// Mitsubishi GX Works2 project: Calculate   PLC: Q06UDEH

TYPE ConveyorIO : STRUCT
  xCWPresent : BOOL;  (* 正转检测有无传感器 *)
  xCCWPresent : BOOL;  (* 反转检测有无传感器 *)
  xLoad : BOOL;  (* 上料请求 *)
  xUnload : BOOL;  (* 下料请求 *)
  xMotorCW : BOOL;  (* 电机正转 *)
  xMotorCCW : BOOL;  (* 电机反转 *)
  xEmpty : BOOL;  (* 线体状态为空 *)
  xNextRun : BOOL;  (* 下段线体运行 *)
  xUnloadCCW : BOOL;  (* 下料为反转 *)
  xloadCCW : BOOL;  (* 上料为反转 *)
  xLeave : BOOL;  (* 已经离开 *)
  xForward : BOOL;  (* 正转手动 *)
  xBackward : BOOL;  (* 反转手动 *)
  xBusy : BOOL;  (* 工作中 *)
  xPutInto : BOOL;  (* 线体直接投入物料 *)
  xLoadAlarrm : BOOL;  (* 上料报警 *)
  xUnloadAlarm : BOOL;  (* 下料报警 *)
  iProductCategory : INT;  (* 产品种类 *)
  tLeaveDelay : TIME;  (* 离开延时设置 *)
  tLoadDelay : TIME;  (* 进入延时设置 *)
END_STRUCT END_TYPE

TYPE ShuttleCarIO : STRUCT
  xReady : BOOL;  (* 准备就绪 *)
  xForward : BOOL;  (* 正转 *)
  xBackward : BOOL;  (* 反转 *)
  iCurrentPos : INT;  (* 当前位置 *)
  iDestinationPos : INT;  (* 目标位置 *)
  xCW : BOOL;  (* 正转输出 *)
  xCCW : BOOL;  (* 反转输出 *)
  xBrake : BOOL;  (* 刹车 *)
  xHomeSwitch : BOOL;  (* 零位接近开关 *)
  xPosLimit : BOOL;  (* 正限位 *)
  xNegLimit : BOOL;  (* 负限位 *)
  xMDIExe : BOOL;  (* MDI开始 *)
  xMDIDone : BOOL;  (* MDI 完成 *)
  xPassLimit : BOOL;  (* 限位屏蔽 *)
  xPosLimitCatch : BOOL;  (* 正限位捕捉 *)
  xNegLimitCatch : BOOL;  (* 负限位捕捉 *)
  xHomeExe : BOOL;  (* 开始寻零 *)
  xHomeDone : BOOL;  (* 寻零完成 *)
  xHomeBusy : BOOL;  (* 寻零中 *)
  xHomeFailed : BOOL;  (* 寻零失败 *)
  xBusy : BOOL;  (* 工作中 *)
END_STRUCT END_TYPE

TYPE SwitchIO : STRUCT
  xLiftCylinderRetractDetect : BOOL;
  xLiftCylinderExtendDetect : BOOL;
  xLiftCylinderRetract : BOOL;
  xLiftCylinderExtend : BOOL;
  xEntryBarCylinderRetract : BOOL;
  xLiftCylinderExtendInit : BOOL;
  xEntryEnable : BOOL;
  xExitEnable : BOOL;
  xExitBarCylinderRetract : BOOL;
  xSwithEnable : BOOL;
  xLiftCylinderRetractButton : BOOL;
  xLiftCylinderExtendButton : BOOL;
  xEntryBarCylinderRetractButton : BOOL;
  xExitBarCylinderRetractButton : BOOL;
END_STRUCT END_TYPE

// global labels: Global1
VAR_GLOBAL
  g_xAuto : BOOL;
  g_xManual : BOOL;
  g_xEStop AT X23 : BOOL;
  g_xReset AT X20 : BOOL;
  g_xStackLampRed AT Y120 : BOOL;
  g_xStackLampAmber AT Y121 : BOOL;
  g_xStackLampGreen AT Y122 : BOOL;
  g_xBuzzer AT Y123 : BOOL;
  g_xStop AT M2 : BOOL;
  g_xLocalAutoStart AT M1 : BOOL;
  g_xRemoteAutoStart AT M0 : BOOL;
  g_xRemoteAuto AT M10 : BOOL;
  g_iState AT D40 : INT;
  g_iLocalAutoStep : INT;
END_VAR

// task Task_01 (event TRUE, interval 0, priority 31): POU, Start, UDP

PROGRAM POU
VAR
  H3000Conveyor1 : Conveyor;
  H3000Conveyor1IO : ConveyorIO;
  H3000Conveyor2 : Conveyor;
  H3000Conveyor2IO : ConveyorIO;
  H3000Conveyor3 : Conveyor;
  H3000Conveyor3IO : ConveyorIO;
  H3000Conveyor4 : Conveyor;
  H3000Conveyor4IO : ConveyorIO;
  H3000Conveyor5 : Conveyor;
  H3000Conveyor5IO : ConveyorIO;
  H3000Conveyor6 : Conveyor;
  H3000Conveyor6IO : ConveyorIO;
  H3000Conveyor7 : Conveyor;
  H3000Conveyor7IO : ConveyorIO;
  H3000Conveyor8 : Conveyor;
  H3000Conveyor8IO : ConveyorIO;
  H3000Conveyor9 : Conveyor;
  H3000Conveyor9IO : ConveyorIO;
  H3000Conveyor10 : Conveyor;
  H3000Conveyor10IO : ConveyorIO;
  H3000ChemConveyor1 : Conveyor;
  H3000ChemConveyor1IO : ConveyorIO;
  H3000ChemConveyor2 : Conveyor;
  H3000ChemConveyor2IO : ConveyorIO;
  H3000ChemConveyor3 : Conveyor;
  H3000ChemConveyor3IO : ConveyorIO;
  Lifter1 : ShuttleCar;
  Lifter1IO : ShuttleCarIO;
  Conveyor1 : Conveyor;
  Conveyor1IO : ConveyorIO;
  Lifter2 : ShuttleCar;
  Lifter2IO : ShuttleCarIO;
  Conveyor2 : Conveyor;
  Conveyor2IO : ConveyorIO;
  H2200Conveyor1 : Conveyor;
  H2200Conveyor1IO : ConveyorIO;
  H2200Conveyor2 : Conveyor;
  H2200Conveyor2IO : ConveyorIO;
  H2200Conveyor3 : Conveyor;
  H2200Conveyor3IO : ConveyorIO;
  H2200Conveyor4 : Conveyor;
  H2200Conveyor4IO : ConveyorIO;
  H2200Conveyor5 : Conveyor;
  H2200Conveyor5IO : ConveyorIO;
  H2200Conveyor6 : Conveyor;
  H2200Conveyor6IO : ConveyorIO;
  H2200Conveyor7 : Conveyor;
  H2200Conveyor7IO : ConveyorIO;
  H2200Conveyor8 : Conveyor;
  H2200Conveyor8IO : ConveyorIO;
  H2200Conveyor9 : Conveyor;
  H2200Conveyor9IO : ConveyorIO;
  H2200Conveyor10 : Conveyor;
  H2200Conveyor10IO : ConveyorIO;
  H1000Conveyor1 : Conveyor;
  H1000Conveyor1IO : ConveyorIO;
  H1000Conveyor2 : Conveyor;
  H1000Conveyor2IO : ConveyorIO;
  H1000Conveyor3 : Conveyor;
  H1000Conveyor3IO : ConveyorIO;
  H1000Conveyor4 : Conveyor;
  H1000Conveyor4IO : ConveyorIO;
  H1000Conveyor5 : Conveyor;
  H1000Conveyor5IO : ConveyorIO;
  H1000Conveyor6 : Conveyor;
  H1000Conveyor6IO : ConveyorIO;
  H1000Conveyor7 : Conveyor;
  H1000Conveyor7IO : ConveyorIO;
  H1000Conveyor8 : Conveyor;
  H1000Conveyor8IO : ConveyorIO;
  H1000Conveyor9 : Conveyor;
  H1000Conveyor9IO : ConveyorIO;
  H3000SwitchChem : Switch;
  H3000SwitchChemIO : SwitchIO;
  H850Switch : Switch;
  H850SwitchIO : SwitchIO;
  H850SwitchConveyorIn : ConveyorIO;
  H850SwitchConveyorOut : ConveyorIO;
  H850Conveyor8 : Conveyor;
  H850Conveyor8IO : ConveyorIO;
  H1000Conveyor10 : Conveyor;
  H1000Conveyor10IO : ConveyorIO;
  H3000SwitchChemConveyorIn : ConveyorIO;
  H3000SwitchChemConveyorOut : ConveyorIO;
  H3000SwitchQuadPackage : Switch;
  H3000SwitchQuadPackageIO : SwitchIO;
  H3000SwitchPackageConveyorIn : ConveyorIO;
  H3000SwitchPackageConveyorOut : ConveyorIO;
  H2200Switch1 : Switch;
  H2200Switch1IO : SwitchIO;
  H2200Switch1ConveyorIn : ConveyorIO;
  H2200Switch1ConveyorOut : ConveyorIO;
  H2200Switch2 : Switch;
  H2200Switch2IO : SwitchIO;
  H2200Switch2ConveyorIn : ConveyorIO;
  H2200Switch2ConveyorOut : ConveyorIO;
  iStep : INT;
  Import1Conveyor1 : Conveyor;
  Import1Conveyor1IO : ConveyorIO;
  Import1Conveyor2 : Conveyor;
  Import1Conveyor2IO : ConveyorIO;
  Import2Conveyor1 : Conveyor;
  Import2Conveyor1IO : ConveyorIO;
  Import2Conveyor2 : Conveyor;
  Import2Conveyor2IO : ConveyorIO;
  Export1Conveyor1 : Conveyor;
  Export1Conveyor1IO : ConveyorIO;
  Export1Conveyor2 : Conveyor;
  Export1Conveyor2IO : ConveyorIO;
  Export2Conveyor1 : Conveyor;
  Export2Conveyor1IO : ConveyorIO;
  Export2Conveyor2 : Conveyor;
  Export2Conveyor2IO : ConveyorIO;
  Export2Switch : Switch;
  Export2SwitchIO : SwitchIO;
  Export2SwitchConveyorIn : ConveyorIO;
  Export2SwitchConveyorOut : ConveyorIO;
  H850Rotor : ShuttleCar;
  H850RotorIO : ShuttleCarIO;
  H850RotorConveyor : Conveyor;
  H850RotorConveyorIO : ConveyorIO;
  H2200RotorIO : ShuttleCarIO;
  H2200RotorConveyor : Conveyor;
  H2200RotorConveyorIO : ConveyorIO;
  H2200Rotor : ShuttleCar;
  H850Conveyor1 : Conveyor;
  H850Conveyor1IO : ConveyorIO;
  H850Conveyor3 : Conveyor;
  H850Conveyor3IO : ConveyorIO;
  H850Conveyor4 : Conveyor;
  H850Conveyor4IO : ConveyorIO;
  H850Conveyor5 : Conveyor;
  H850Conveyor5IO : ConveyorIO;
  H850Conveyor6 : Conveyor;
  H850Conveyor6IO : ConveyorIO;
  Lifter2Position : ARRAY [0..5] OF INT;
  ii : INT;
  H2200SwitchEmptyABack : Switch;
  H2200SwitchEmptyABackIO : SwitchIO;
  H2200SwitchEmptyABackConveyorIn : ConveyorIO;
  H2200SwitchEmptyABackConveyorOut : ConveyorIO;
  H2200SwitchEmptyBBack : Switch;
  H2200SwitchEmptyBBackIO : SwitchIO;
  H2200SwitchEmptyBBackConveyorIn : ConveyorIO;
  H2200SwitchEmptyBBackConveyorOut : ConveyorIO;
  H2200ImportConveyor1 : Conveyor;
  H2200ImportConveyor1IO : ConveyorIO;
  H2200ImportConveyor2 : Conveyor;
  H2200ImportConveyor2IO : ConveyorIO;
  Import1Switch : Switch;
  Import1SwitchIO : SwitchIO;
  Import1SwitchConveyorIn : ConveyorIO;
  Import1SwitchConveyorOut : ConveyorIO;
  Export1Switch : Switch;
  Export1SwitchIO : SwitchIO;
  Export1SwitchConveyorIn : ConveyorIO;
  Export1SwitchConveyorOut : ConveyorIO;
  Import2Switch : Switch;
  Import2SwitchIO : SwitchIO;
  Import2SwitchConveyorIn : ConveyorIO;
  Import2SwitchConveyorOut : ConveyorIO;
  Import1LoadCylinder : ShuttleCar;
  Import1LoadCylinderIO : ShuttleCarIO;
  Import2LoadCylinder : ShuttleCar;
  Import2LoadCylinderIO : ShuttleCarIO;
  Export1LoadCylinder : ShuttleCar;
  Export1LoadCylinderIO : ShuttleCarIO;
  Export2LoadCylinder : ShuttleCar;
  Export2LoadCylinderIO : ShuttleCarIO;
  Lifter2Occupy : BOOL;  (* 提升机2占用标志位 *)
  Lifter2ChemImport : BOOL;  (* 提升机2化成入库 *)
  Lifter2ExportChem : BOOL;  (* 提升机2出库到化成 *)
END_VAR
H3000SwitchQuadPackage(ConveyorEntryIO:=H3000SwitchPackageConveyorIn ,
                                                        ConveyorExitIO:=H3000SwitchPackageConveyorOut ,
                                                        SwitchIO:=H3000SwitchQuadPackageIO );
H3000SwitchQuadPackageIO.xLiftCylinderExtendButton:=M75;
H3000SwitchQuadPackageIO.xLiftCylinderRetractButton:=M76;
H3000SwitchQuadPackageIO.xExitBarCylinderRetractButton:=M83;
Y128:=H3000SwitchQuadPackageIO.xEXITBarCylinderRetract;
Y12C:=H3000SwitchQuadPackageIO.xLiftCylinderExtend;
Y12A:=H3000SwitchQuadPackageIO.xLiftCylinderRetract;
H3000SwitchQuadPackageIO.xLiftCylinderExtendDetect:=X29;
H3000SwitchQuadPackageIO.xLiftCylinderRetractDetect:=X2A;
H3000SwitchPackageConveyorIn.xForward:=M77;
H3000SwitchPackageConveyorIn.xCWPresent:=X28;
(*Y187:=H3000SwitchPackageConveyorIn.xMotorCW;*)
H3000SwitchPackageConveyorOut.xForward:=M78;
H3000SwitchPackageConveyorOut.xCWPresent:=X2B;
Y12B:=H3000SwitchPackageConveyorOut.xMotorCW;

H3000SwitchChem(ConveyorEntryIO:=H3000SwitchChemConveyorIn ,
                                                        ConveyorExitIO:=H3000SwitchChemConveyorOut ,
                                                        SwitchIO:=H3000SwitchChemIO );
H3000SwitchChemIO.xLiftCylinderExtendButton:=M79;
H3000SwitchChemIO.xLiftCylinderRetractButton:=M80;
Y129:=H3000SwitchChemIO.xLiftCylinderExtend;
Y12D:=H3000SwitchChemIO.xLiftCylinderRetract;
H3000SwitchChemIO.xLiftCylinderExtendDetect:=X2C;
H3000SwitchChemIO.xLiftCylinderRetractDetect:=X2D;
H3000SwitchChemConveyorIn.xForward:=M81;
H3000SwitchChemConveyorIn.xCWPresent:=X2E;
Y19B:=H3000SwitchPackageConveyorIn.xMotorCW;
H3000SwitchChemConveyorOut.xForward:=M82;
H3000SwitchChemConveyorOut.xCWPresent:=X2E;
Y12E:=H3000SwitchChemConveyorOut.xMotorCW;
H3000SwitchChemIO.xSwithEnable:=1;

Lifter1(ShuttleCarInOut:=Lifter1IO);
ShuttleCarCurrentPosition( X8C OR X8D ,X8C ,X8D, FALSE, Lifter1IO.iCurrentPos );
Lifter1IO.xReady:=X24;
Lifter1Io.xForward:=M50 OR X91;
Lifter1IO.xBackward:=M51 OR X92;
Lifter1IO.xPosLimit:=X8E;
Lifter1IO.xNegLimit:=X8F;
Y18D:=Lifter1IO.xCW;
Y18E:=Lifter1IO.xCCW;
Y192:=Lifter1IO.xBrake;

Conveyor1(ConveyorMotor:=Conveyor1IO);
Conveyor1IO.xForward:=M52;
Conveyor1IO.xBackward:=M53;
Conveyor1IO.xCWPresent:=X93;
Conveyor1IO.xCCWPresent:=X94;
Y18B:=Conveyor1IO.xMotorCW;
Y18C:=Conveyor1IO.xMotorCCW;

Lifter2(ShuttleCarInOut:=Lifter2IO);
Lifter2Position[0]:=0;
Lifter2Position[1]:=57;
Lifter2Position[2]:=590;
Lifter2Position[3]:=5828;
Lifter2Position[4]:=6202;
Lifter2Position[5]:=9200;
FOR ii:=0 TO 5 BY 1 DO
	IF abs(D190-Lifter2Position[ii])<5 THEN
		Lifter2IO.iCurrentPos:=ii;
	END_IF;
END_FOR;
Lifter2IO.xReady:=X25;
(*提升机占用标志位控制*)
IF LIfter2IO.xBusy AND Conveyor2IO.xEmpty=0 AND g_xAuto THEN
	Lifter2Occupy:=1;
END_IF;
IF g_xManual OR g_xReset THEN
	Lifter2Occupy:=0;
END_IF;
IF ( Lifter2IO.iCurrentPos=1 AND NOT H850Conveyor8IO.xEmpty)   (*注液入库*)
	OR (Lifter2IO.iCurrentPos=2 AND NOT H1000Conveyor1IO.xEmpty)  (*化成入库*)
	OR (Lifter2IO.iCurrentPos=5  AND NOT H3000ChemConveyor3IO.xEmpty) THEN(*出库化成或空框去注液*)
	Lifter2Occupy:=1;
END_IF;
IF  (Lifter2IO.iCurrentPos=3 OR Lifter2IO.iCurrentPos=4) AND Conveyor2IO.xEmpty  THEN
	Lifter2Occupy:=0;
END_IF;

Lifter2Io.xForward:=M54 OR X9B;
Lifter2IO.xBackward:=M55 OR X9C;
Lifter2IO.xPosLimit:=X98;
Lifter2IO.xNegLimit:=X99;
Y193:=Lifter2IO.xCW;
Y194:=Lifter2IO.xCCW;
Y198:=Lifter2IO.xBrake;
(*提升机2编码器清零，到达负限位后清零*)
IF NOT Lifter2IO.xNegLimit THEN
	Y125:=1;
ELSE
	Y125:=0;
END_IF;

Conveyor2(ConveyorMotor:=Conveyor2IO);
Conveyor2IO.xForward:=M56;
Conveyor2IO.xBackward:=M57;
Conveyor2IO.xCWPresent:=X9D;
Conveyor2IO.xCCWPresent:=X9E;
Y19A:=Conveyor2IO.xMotorCW;
Y199:=Conveyor2IO.xMotorCCW;


H3000Conveyor1(ConveyorMotor:=H3000Conveyor1IO);
H3000Conveyor1IO.xForward:=M30;
H3000Conveyor1IO.xCWPresent:=X2F;
Y12F:=H3000Conveyor1IO.xMotorCW;

H3000Conveyor2(ConveyorMotor:=H3000Conveyor2IO);
H3000Conveyor2IO.xForward:=M31;
H3000Conveyor2IO.xCWPresent:=X30;
Y130:=H3000Conveyor2IO.xMotorCW;

H3000Conveyor3(ConveyorMotor:=H3000Conveyor3IO);
H3000Conveyor3IO.xForward:=M32;
H3000Conveyor3IO.xCWPresent:=X31;
Y131:=H3000Conveyor3IO.xMotorCW;

H3000Conveyor4(ConveyorMotor:=H3000Conveyor4IO);
H3000Conveyor4IO.xForward:=M33;
H3000Conveyor4IO.xCWPresent:=X32;
Y132:=H3000Conveyor4IO.xMotorCW;

H3000Conveyor5(ConveyorMotor:=H3000Conveyor5IO);
H3000Conveyor5IO.xForward:=M34;
H3000Conveyor5IO.xCWPresent:=X33;
Y133:=H3000Conveyor5IO.xMotorCW;

H3000Conveyor6(ConveyorMotor:=H3000Conveyor6IO);
H3000Conveyor6IO.xForward:=M34;
H3000Conveyor6IO.xCWPresent:=X34;
Y134:=H3000Conveyor6IO.xMotorCW;

H3000Conveyor7(ConveyorMotor:=H3000Conveyor7IO);
H3000Conveyor7IO.xForward:=M35;
H3000Conveyor7IO.xCWPresent:=X35;
Y135:=H3000Conveyor7IO.xMotorCW;
H3000Conveyor8(ConveyorMotor:=H3000Conveyor8IO);
H3000Conveyor8IO.xForward:=M36;
H3000Conveyor8IO.xCWPresent:=X36;
Y136:=H3000Conveyor8IO.xMotorCW;

H3000Conveyor9(ConveyorMotor:=H3000Conveyor9IO);
H3000Conveyor9IO.xForward:=M37;
H3000Conveyor9IO.xCWPresent:=X37;
Y137:=H3000Conveyor9IO.xMotorCW;

H3000Conveyor10(ConveyorMotor:=H3000Conveyor10IO);
H3000Conveyor10IO.xForward:=M38;
H3000Conveyor10IO.xCWPresent:=X38;
Y138:=H3000Conveyor10IO.xMotorCW;

H3000ChemConveyor1(ConveyorMotor:=H3000ChemConveyor1IO);
H3000ChemConveyor1IO.xForward:=M39;
H3000ChemConveyor1IO.xCWPresent:=X39;
Y139:=H3000ChemConveyor1IO.xMotorCW;

H3000ChemConveyor2(ConveyorMotor:=H3000ChemConveyor2IO);
H3000ChemConveyor2IO.xForward:=M40;
H3000ChemConveyor2IO.xCWPresent:=X3A;
Y13A:=H3000ChemConveyor2IO.xMotorCW;

H3000ChemConveyor3(ConveyorMotor:=H3000ChemConveyor3IO);
H3000ChemConveyor3IO.xForward:=M41;
H3000ChemConveyor3IO.xCWPresent:=X3B;
Y13B:=H3000ChemConveyor3IO.xMotorCW;

H2200Switch1(ConveyorEntryIO:=H2200Switch1ConveyorIn ,
                                                        ConveyorExitIO:=H2200Switch1ConveyorOut ,
                                                        SwitchIO:=H2200Switch1IO );
H2200Switch1IO.xLiftCylinderExtendButton:=M84;
H2200Switch1IO.xLiftCylinderRetractButton:=M85;
H2200Switch1IO.xExitBarCylinderRetractButton:=M86;
Y158:=H2200Switch1IO.xEXITBarCylinderRetract;
Y155:=H2200Switch1IO.xLiftCylinderExtend;
Y156:=H2200Switch1IO.xLiftCylinderRetract;
H2200Switch1IO.xLiftCylinderExtendDetect:=X55;
H2200Switch1IO.xLiftCylinderRetractDetect:=X56;
H2200Switch1ConveyorIn.xForward:=M87;
H2200Switch1ConveyorIn.xCWPresent:=X57;
Y177:=H2200Switch1ConveyorIn.xMotorCW;
H2200Switch1ConveyorOut .xForward:=M88;
H2200Switch1ConveyorOut .xCWPresent:=X57;
H2200Switch1ConveyorOut.tLoadDelay:=T#1s;
Y157:=H2200Switch1ConveyorOut .xMotorCW;

H2200ImportConveyor1(ConveyorMotor:=H2200ImportConveyor1IO);
H2200ImportConveyor1IO.xForward:=M136;
H2200ImportConveyor1IO.xCWPresent:=X53;
Y153:=H2200ImportConveyor1IO.xMotorCW;
H2200ImportConveyor2IO.tLeaveDelay:=T#5s;

H2200ImportConveyor2(ConveyorMotor:=H2200ImportConveyor2IO);
H2200ImportConveyor2IO.xForward:=M122;
H2200ImportConveyor2IO.xCWPresent:=X58;
Y154:=H2200ImportConveyor2IO.xMotorCW;
H2200ImportConveyor2IO.tLeaveDelay:=T#5s;

H2200Switch2(ConveyorEntryIO:=H2200Switch2ConveyorIn ,
                                                        ConveyorExitIO:=H2200Switch2ConveyorOut ,
                                                        SwitchIO:=H2200Switch2IO );
H2200Switch2IO.xLiftCylinderExtendButton:=M89;
H2200Switch2IO.xLiftCylinderRetractButton:=M90;
H2200Switch2IO.xExitBarCylinderRetractButton:=M91;
Y15C:=H2200Switch2IO.xEXITBarCylinderRetract;
Y159:=H2200Switch2IO.xLiftCylinderExtend;
Y15A:=H2200Switch2IO.xLiftCylinderRetract;
H2200Switch2IO.xLiftCylinderExtendDetect:=X59;
H2200Switch2IO.xLiftCylinderRetractDetect:=X5A;
H2200Switch2ConveyorIn.xForward:=M92;
H2200Switch2ConveyorIn.xCWPresent:=X5B;
H2200Switch2ConveyorIn.tLoadDelay:=T#2s;
Y15B:=H2200Switch2ConveyorIn.xMotorCW;
H2200Switch2ConveyorOut .xForward:=M93;
H2200Switch2ConveyorOut .xCWPresent:=X5B;
H2200Switch2ConveyorOut.tLeaveDelay:=T#8S;
H2200Switch2IO.xLiftCylinderExtendInit:=1;

H2200SwitchEmptyABack(ConveyorEntryIO:=H2200SwitchEmptyABackConveyorIn ,
                                                        ConveyorExitIO:=H2200SwitchEmptyABackConveyorOut ,
                                                        SwitchIO:=H2200SwitchEmptyABackIO );
H2200SwitchEmptyABackIO.xLiftCylinderExtendButton:=M137;
H2200SwitchEmptyABackIO.xLiftCylinderRetractButton:=M138;
H2200SwitchEmptyABackIO.xExitBarCylinderRetractButton:=M139;
Y160:=H2200SwitchEmptyABackIO.xLiftCylinderExtend;
Y161:=H2200SwitchEmptyABackIO.xLiftCylinderRetract;
H2200SwitchEmptyABackIO.xLiftCylinderExtendDetect:=X60;
H2200SwitchEmptyABackIO.xLiftCylinderRetractDetect:=X61;
H2200SwitchEmptyABackConveyorIn.xForward:=M140;
H2200SwitchEmptyABackConveyorIn.xCWPresent:=X62;
H2200SwitchEmptyABackConveyorIn.tLoadDelay:=T#2s;
Y162:=H2200SwitchEmptyABackConveyorIn.xMotorCW;
H2200SwitchEmptyABackConveyorOut .xForward:=M146;
H2200SwitchEmptyABackConveyorOut.xCWPresent:=X62;
H2200SwitchEmptyABackConveyorOut.tLeaveDelay:=T#30S;
Y177:=H2200SwitchEmptyABackConveyorOut .xMotorCW OR H2200SwitchEmptyBBackConveyorOut .xMotorCW ;

H2200SwitchEmptyBBack(ConveyorEntryIO:=H2200SwitchEmptyBBackConveyorIn ,
                                                        ConveyorExitIO:=H2200SwitchEmptyBBackConveyorOut ,
                                                        SwitchIO:=H2200SwitchEmptyBBackIO );
H2200SwitchEmptyBBackIO.xLiftCylinderExtendButton:=M141;
H2200SwitchEmptyBBackIO.xLiftCylinderRetractButton:=M142;
H2200SwitchEmptyBBackIO.xExitBarCylinderRetractButton:=M143;
Y166:=H2200SwitchEmptyBBackIO.xLiftCylinderExtend;
Y167:=H2200SwitchEmptyBBackIO.xLiftCylinderRetract;
H2200SwitchEmptyBBackIO.xLiftCylinderExtendDetect:=X66;
H2200SwitchEmptyBBackIO.xLiftCylinderRetractDetect:=X67;
H2200SwitchEmptyBBackConveyorIn.xForward:=M144;
H2200SwitchEmptyBBackConveyorIn.xCWPresent:=X68;
H2200SwitchEmptyBBackConveyorIn.tLoadDelay:=T#2s;
Y168:=H2200SwitchEmptyBBackConveyorIn.xMotorCW;
H2200SwitchEmptyBBackConveyorOut .xForward:=M145;
H2200SwitchEmptyBBackConveyorOut.xCWPresent:=X68;
H2200SwitchEmptyBBackConveyorOut.tLeaveDelay:=T#30S;

H2200Rotor(ShuttleCarInOut:=H2200RotorIO);
ShuttleCarCurrentPosition( X6F OR X75 ,X6F ,X75, FALSE, H2200RotorIO.iCurrentPos );
H2200RotorIO.xReady:=TRUE;
H2200RotorIO.xForward:=M78;
H2200RotorIO.xBackward:=M79;
H2200RotorIO.xPosLimit:=X71;
H2200RotorIO.xNegLimit:=X72;
Y170:=H2200RotorIO.xCW;
Y16F:=H2200RotorIO.xCCW;
Y1B8:=H2200RotorIO.xBrake;

H2200RotorConveyor(ConveyorMotor:=H2200RotorConveyorIO);
H2200RotorConveyorIO.xForward:=M80;
H2200RotorConveyorIO.xBackward:=M81;
H2200RotorConveyorIO.xCWPresent:=X74;
H2200RotorConveyorIO.xCcWPresent:=X73;
Y172:=H2200RotorConveyorIO.xMotorCW;
Y171:=H2200RotorConveyorIO.xMotorCCW;

H2200Conveyor1(ConveyorMotor:=H2200Conveyor1IO);
H2200Conveyor1IO.xForward:=M42;
H2200Conveyor1IO.xCWPresent:=X3F;
Y13F:=H2200Conveyor1IO.xMotorCW;

H2200Conveyor2(ConveyorMotor:=H2200Conveyor2IO);
H2200Conveyor2IO.xForward:=M43;
H2200Conveyor2IO.xCWPresent:=X40;
Y140:=H2200Conveyor2IO.xMotorCW;

H2200Conveyor3(ConveyorMotor:=H2200Conveyor3IO);
H2200Conveyor3IO.xForward:=M44;
H2200Conveyor3IO.xCWPresent:=X41;
Y141:=H2200Conveyor3IO.xMotorCW;

H2200Conveyor4(ConveyorMotor:=H2200Conveyor4IO);
H2200Conveyor4IO.xForward:=M45;
H2200Conveyor4IO.xCWPresent:=X42;
Y142:=H2200Conveyor4IO.xMotorCW;

H2200Conveyor5(ConveyorMotor:=H2200Conveyor5IO);
H2200Conveyor5IO.xForward:=M46;
H2200Conveyor5IO.xCWPresent:=X43;
Y143:=H2200Conveyor5IO.xMotorCW;

H2200Conveyor6(ConveyorMotor:=H2200Conveyor6IO);
H2200Conveyor6IO.xForward:=M47;
H2200Conveyor6IO.xCWPresent:=X44;
Y144:=H2200Conveyor6IO.xMotorCW;

H2200Conveyor7(ConveyorMotor:=H2200Conveyor7IO);
H2200Conveyor7IO.xForward:=M48;
H2200Conveyor7IO.xCWPresent:=X45;
Y145:=H2200Conveyor7IO.xMotorCW;

H2200Conveyor8(ConveyorMotor:=H2200Conveyor8IO);
H2200Conveyor8IO.xForward:=M49;
H2200Conveyor8IO.xCWPresent:=X46;
Y146:=H2200Conveyor8IO.xMotorCW;

H2200Conveyor9(ConveyorMotor:=H2200Conveyor9IO);
H2200Conveyor9IO.xForward:=M58;
H2200Conveyor9IO.xCWPresent:=X47;
Y147:=H2200Conveyor9IO.xMotorCW;

H2200Conveyor10(ConveyorMotor:=H2200Conveyor10IO);
H2200Conveyor10IO.xForward:=M59;
H2200Conveyor10IO.xCWPresent:=X48;
Y148:=H2200Conveyor10IO.xMotorCW;

H1000Conveyor1(ConveyorMotor:=H1000Conveyor1IO);
H1000Conveyor1IO.xForward:=M60;
H1000Conveyor1IO.xCWPresent:=X49;
Y149:=H1000Conveyor1IO.xMotorCW;

H1000Conveyor2(ConveyorMotor:=H1000Conveyor2IO);
H1000Conveyor2IO.xForward:=M61;
H1000Conveyor2IO.xCWPresent:=X4A;
Y14A:=H1000Conveyor2IO.xMotorCW;

H1000Conveyor3(ConveyorMotor:=H1000Conveyor3IO);
H1000Conveyor3IO.xForward:=M62;
H1000Conveyor3IO.xCWPresent:=X4B;
Y14B:=H1000Conveyor3IO.xMotorCW;

H1000Conveyor4(ConveyorMotor:=H1000Conveyor4IO);
H1000Conveyor4IO.xForward:=M63;
H1000Conveyor4IO.xCWPresent:=X4C;
Y14C:=H1000Conveyor4IO.xMotorCW;

H1000Conveyor5(ConveyorMotor:=H1000Conveyor5IO);
H1000Conveyor5IO.xForward:=M64;
H1000Conveyor5IO.xCWPresent:=X4D;
Y14D:=H1000Conveyor5IO.xMotorCW;

H1000Conveyor6(ConveyorMotor:=H1000Conveyor6IO);
H1000Conveyor6IO.xForward:=M65;
H1000Conveyor6IO.xCWPresent:=X4E;
Y14E:=H1000Conveyor6IO.xMotorCW;

H1000Conveyor7(ConveyorMotor:=H1000Conveyor7IO);
H1000Conveyor7IO.xForward:=M66;
H1000Conveyor7IO.xCWPresent:=X4F;
Y14F:=H1000Conveyor7IO.xMotorCW;

H1000Conveyor8(ConveyorMotor:=H1000Conveyor8IO);
H1000Conveyor8IO.xForward:=M67;
H1000Conveyor8IO.xCWPresent:=X50;
Y150:=H1000Conveyor8IO.xMotorCW;

H1000Conveyor9(ConveyorMotor:=H1000Conveyor9IO);
H1000Conveyor9IO.xForward:=M68;
H1000Conveyor9IO.xCWPresent:=X51;
Y151:=H1000Conveyor9IO.xMotorCW;

H1000Conveyor10(ConveyorMotor:=H1000Conveyor10IO);
H1000Conveyor10IO.xForward:=M67;
H1000Conveyor10IO.xCWPresent:=X52;
Y152:=H1000Conveyor10IO.xMotorCW;

H850Conveyor1(ConveyorMotor:=H850Conveyor1IO);
H850Conveyor1IO.xForward:=M129;
H850Conveyor1IO.xCWPresent:=X78;
Y178:=H850Conveyor1IO.xMotorCW;

H850Conveyor3(ConveyorMotor:=H850Conveyor3IO);
H850Conveyor3IO.xForward:=M130;
H850Conveyor3IO.xCWPresent:=X7A;
Y17A:=H850Conveyor3IO.xMotorCW;

H850Conveyor4(ConveyorMotor:=H850Conveyor4IO);
H850Conveyor4IO.xForward:=M131;
H850Conveyor4IO.xCWPresent:=X7B;
Y17B:=H850Conveyor4IO.xMotorCW;

H850Conveyor5(ConveyorMotor:=H850Conveyor5IO);
H850Conveyor5IO.xForward:=M132;
H850Conveyor5IO.xCWPresent:=X7C;
Y17C:=H850Conveyor5IO.xMotorCW;

H850Conveyor6(ConveyorMotor:=H850Conveyor6IO);
H850Conveyor6IO.xForward:=M133;
H850Conveyor6IO.xCWPresent:=X7D;
Y17D:=H850Conveyor6IO.xMotorCW;

H850Rotor(ShuttleCarInOut:=H850RotorIO);
ShuttleCarCurrentPosition( X82 OR X76 ,X82 ,X76, FALSE, H850RotorIO.iCurrentPos );
H850RotorIO.xReady:=TRUE;
H850RotorIO.xForward:=M75;
H850RotorIO.xBackward:=M76;
H850RotorIO.xPosLimit:=X84;
H850RotorIO.xNegLimit:=X85;
Y182:=H850RotorIO.xCW;
Y183:=H850RotorIO.xCCW;
Y1B9:=H850RotorIO.xBrake;

H850RotorConveyor(ConveyorMotor:=H850RotorConveyorIO);
H850RotorConveyorIO.xForward:=M77;
H850RotorConveyorIO.xBackward:=M82;
H850RotorConveyorIO.xCWPresent:=X87;
H850RotorConveyorIO.xCCWPresent:=X86;
Y185:=H850RotorConveyorIO.xMotorCW;
Y184:=H850RotorConveyorIO.xMotorCCW;
H850RotorConveyorIO.xUnloadCCW:=1;
H850RotorConveyorIO.tLeaveDelay:=T#10s;

H850Switch(ConveyorEntryIO:=H850SwitchConveyorIn,ConveyorExitIO:=H850SwitchConveyorOut,SwitchIO:=H850SwitchIO);
H850SwitchIO.xLiftCylinderExtendButton:=M71;
H850SwitchIO.xLiftCylinderRetractButton:=M72;
Y189:=H850SwitchIO.xLiftCylinderExtend;
Y188:=H850SwitchIO.xLiftCylinderRetract;
H850SwitchIO.xLiftCylinderExtendDetect:=X88;
H850SwitchIO.xLiftCylinderRetractDetect:=X89;
H850SwitchConveyorIn.xForward:=M70;
H850SwitchConveyorIn.xCWPresent:=XB4;
Y19B:=H850SwitchConveyorIn.xMotorCW;
H850SwitchConveyorOut.xForward:=M73;
H850SwitchConveyorOut.xCWPresent:=X8A;
H850SwitchConveyorOut.tLeaveDelay:=T#10s;
Y18A:=H850SwitchConveyorOut.xMotorCW;


H850Conveyor8(ConveyorMotor:=H850Conveyor8IO);
H850Conveyor8IO.xForward:=M74;
H850Conveyor8IO.xCWPresent:=X7F;
Y17F:=H850Conveyor8IO.xMotorCW;
H850Conveyor8IO.tLeaveDelay:=T#5s;

(*高温库前线体*)
(*1巷道入库*)
Import1Conveyor1(ConveyorMotor:=Import1Conveyor1IO);
Import1Conveyor1IO.tLeaveDelay:=t#10s;
Import1Conveyor1IO.xForward:=M98;
Import1Conveyor1IO.xCWPresent:=XE3;
Y1F4:=Import1Conveyor1IO.xMotorCW;

Import1Conveyor2(ConveyorMotor:=Import1Conveyor2IO);
Import1Conveyor2IO.tLeaveDelay:=t#10s;
Import1Conveyor2IO.xForward:=M99;
Import1Conveyor2IO.xCWPresent:=XE4;
Y1F5:=Import1Conveyor2IO.xMotorCW;

Import1Switch(ConveyorEntryIO:=Import1SwitchConveyorIn,
                          ConveyorExitIO:=Import1SwitchConveyorOut ,
                           SwitchIO:=Import1SwitchIO);
Import1SwitchIO.xLiftCylinderExtendButton:=M147;
Import1SwitchIO.xLiftCylinderRetractButton:=M148;
Import1SwitchIO.xExitBarCylinderRetractButton:=M161;
Y1E0:=Import1SwitchIO.xExitBarCylinderRetract;
Y1E2:=Import1SwitchIO.xLiftCylinderExtend;
Y1E1:=Import1SwitchIO.xLiftCylinderRetract;
Import1SwitchIO.xLiftCylinderExtendDetect:=XE1;
Import1SwitchIO.xLiftCylinderRetractDetect:=XE2;
Import1SwitchConveyorIn.xCWPresent:=XE0;
Import1SwitchConveyorIn.tLoadDelay:=T#2s;
Import1SwitchConveyorOut.xForward:=M149;
Import1SwitchConveyorOut.xCWPresent:=X108;
Import1SwitchConveyorOut.tLeaveDelay:=t#8s;
Y1F6:=Import1SwitchConveyorOut.xMotorCW;

Import1LoadCylinder(ShuttleCarInOut:=Import1LoadCylinderIO);
ShuttleCarCurrentPosition( XE6 OR XE7 ,XE7 ,XE6, FALSE, Import1LoadCylinderIO.iCurrentPos );
Import1LoadCylinderIO.xReady:=TRUE;
Import1LoadCylinderIO.xForward:=M159;
Import1LoadCylinderIO.xBackward:=M160;
Import1LoadCylinderIO.xPosLimit:=TRUE;
Import1LoadCylinderIO.xNegLimit:=TRUE;
Y1E4:=Import1LoadCylinderIO.xCW;
Y1E3:=Import1LoadCylinderIO.xCCW;

(*1巷道出库*)
Export1Conveyor1(ConveyorMotor:=Export1Conveyor1IO);
Export1Conveyor1IO.tLeaveDelay:=t#10s;
Export1Conveyor1IO.xForward:=M94;
Export1Conveyor1IO.xCWPresent:=XEB;
Y1F7:=Export1Conveyor1IO.xMotorCW;

Export1Conveyor2(ConveyorMotor:=Export1Conveyor2iO);
Export1Conveyor2IO.tLeaveDelay:=t#10s;
Export1Conveyor2IO.xForward:=M95;
Export1Conveyor2IO.xCWPresent:=XEC;
Y1F8:=Export1Conveyor2IO.xMotorCW;

Export1Switch(ConveyorEntryIO:=Export1SwitchConveyorIn,
                          ConveyorExitIO:=Export1SwitchConveyorOut ,
                           SwitchIO:=Export1SwitchIO);
Export1SwitchIO.xLiftCylinderExtendButton:=M150;
Export1SwitchIO.xLiftCylinderRetractButton:=M151;
Y1E7:=Export1SwitchIO.xLiftCylinderExtend;
Y1E6:=Export1SwitchIO.xLiftCylinderRetract;
Export1SwitchIO.xLiftCylinderExtendDetect:=XE9;
Export1SwitchIO.xLiftCylinderRetractDetect:=XEA;
Export1SwitchConveyorIn.xForward:=M152;
Export1SwitchConveyorIn.xCWPresent:=X106;
Export1SwitchConveyorIn.tLoadDelay:=T#2s;
Y1FF:=Export1SwitchConveyorIn.xMotorCW;
Export1SwitchConveyorOut.xCWPresent:=X106;

Export1LoadCylinder(ShuttleCarInOut:=Export1LoadCylinderIO);
ShuttleCarCurrentPosition( XEF OR XEE ,XEF ,XEE, FALSE, Export1LoadCylinderIO.iCurrentPos );
Export1LoadCylinderIO.xReady:=TRUE;
Export1LoadCylinderIO.xForward:=M157;
Export1LoadCylinderIO.xBackward:=M158;
Export1LoadCylinderIO.xPosLimit:=TRUE;
Export1LoadCylinderIO.xNegLimit:=TRUE;
Y1E8:=Export1LoadCylinderIO.xCW;
Y1E9:=Export1LoadCylinderIO.xCCW;


(*2巷道入库*)
Import2Conveyor1(ConveyorMotor:=Import2Conveyor1IO);
Import2Conveyor1IO.tLeaveDelay:=t#10s;
Import2Conveyor1IO.xForward:=M153;
Import2Conveyor1IO.xCWPresent:=XF3;
Y1FA:=Import2Conveyor1IO.xMotorCW;

Import2Conveyor2(ConveyorMotor:=Import2Conveyor1IO);
Import2Conveyor2IO.tLeaveDelay:=t#10s;
Import2Conveyor2IO.xForward:=M154;
Import2Conveyor2IO.xCWPresent:=XF4;
Y1FB:=Import2Conveyor2IO.xMotorCW;